// TIA Portal project "SSA-3GHz" (V15.1)

(* hardware
DEVICE "S7-1200"  S7-1200 Station
   slot 0: "Stand.sectionalRail35mmLength483mm_0"  S7-1200 Rack  Rack  V1.0
   slot 1: "S7-1200"  CPU 1215C DC/DC/DC  6ES7 215-1AG40-0XB0  V4.3
   slot 2: "AnalogInputSM12314AI_2"  6ES7 231-4HD32-0XB0  V2.0
   slot 3: "S7-1200analogInputSM1231RTD4AI_3"  SM 1231 AI4 x RTD  6ES7 231-5PD32-0XB0  V2.0
DEVICE "HMI_1"  KTP400 Basic PN
   slot 0: "HMI_1"  KTP400 Basic PN  6AV2 123-2DB03-0AX0  15.1.0.0
   slot 1: "HMI_RT_1"  KTP400 Basic PN  6AV2 123-2DB03-0AX0  15.1.0.0
   slot 5: "HMI_1.IE_CP_1"  PROFINET Interface  15.0.1.0
      slot 1: "PROFINET Interface_1"  PROFINET Interface
         slot 1: "Port_1"  Port
*)

// ===== PLC "S7-1200"  CPU 1215C DC/DC/DC =====

VAR_GLOBAL   // PLC tag table "Default tag table"
   "System_Byte" AT %MB1 : Byte;
   "FirstScan" AT %M1.0 : Bool;
   "DiagStatusUpdate" AT %M1.1 : Bool;
   "AlwaysTRUE" AT %M1.2 : Bool;
   "AlwaysFALSE" AT %M1.3 : Bool;
   "Clock_Byte" AT %MB0 : Byte;
   "Clock_10Hz" AT %M0.0 : Bool;
   "Clock_5Hz" AT %M0.1 : Bool;
   "Clock_2.5Hz" AT %M0.2 : Bool;
   "Clock_2Hz" AT %M0.3 : Bool;
   "Clock_1.25Hz" AT %M0.4 : Bool;
   "Clock_1Hz" AT %M0.5 : Bool;
   "Clock_0.625Hz" AT %M0.6 : Bool;
   "Clock_0.5Hz" AT %M0.7 : Bool;
   "MoveBlkStat" AT %MW100 : Int;
END_VAR

VAR_GLOBAL   // PLC tag table "Test tags"
   "Counter" AT %MD100 : UDInt;
   "TestBlink" AT %Q1.0 : Bool;
   "VisuTest" AT %MB104 : Byte;
END_VAR

VAR_GLOBAL   // PLC tag table "Analog I/O"
   "U_drain_RBK" AT %IW64 : Int;   // Drain voltage read-back
   "U_drain" AT %QW64 : Int;   // Drain voltage set-point
   "ADC0ch1" AT %IW66 : Int;   // Spare
   "U_gate" AT %QW66 : Int;   // Gate voltage set-point
   "Pfwd" AT %IW96 : Int;   // Forward power
   "Prev" AT %IW98 : Int;   // Reverse power
   "I_drain" AT %IW100 : Int;   // Drain current
   "U_gate_RBK" AT %IW102 : Int;   // Gate voltage read-back
   "TT001" AT %IW112 : Int;
   "TT002" AT %IW114 : Int;
   "TT003" AT %IW116 : Int;
   "TT004" AT %IW118 : Int;
END_VAR

VAR_GLOBAL   // PLC tag table "Digital I/O"
   "DutyCycOK" AT %I0.0 : Bool;   // Duty cycle OK
   "KeyIntlkOK" AT %I0.1 : Bool;   // Key interlock OK
   "ExtIntlkT1" AT %I0.2 : Bool;   // DC PS enable
   "ExtIntlkT3" AT %I0.3 : Bool;
   "PS_OK" AT %I0.4 : Bool;
   "CoolingWtrOK" AT %I0.5 : Bool;
   "KeyOK" AT %I0.6 : Bool;
   "FanOK" AT %I0.7 : Bool;
   "ExtIntlkOK" AT %I1.0 : Bool;
   "RFSwitchOn" AT %Q0.0 : Bool;   // Close RF switch
   "PScmdOn" AT %Q0.1 : Bool;   // Set PS On
   "SSA_OK" AT %Q0.2 : Bool;   // Solid State Amplifier OK
   "ResetOut" AT %Q0.3 : Bool;   // Reset the errors signal out
END_VAR

TYPE "DigitalIN"
   STRUCT
      DigitalIN : Struct
         PhysIn : Bool;   // Physical input
         NegLogic : Bool;   // 0 - positive lgic, 1 - negative logic
         Disabled : Bool;   // 0 - signal enabled, 1 - signal disabled (not used in process controll)
         Out : Bool;   // Logical value after taking into accout NegLogic setting
      END_STRUCT;
   END_STRUCT;
END_TYPE

TYPE "AnalogOUT"
   STRUCT
      AnalogOUT : Struct
         In : Real;
         Out : Int;
         VisuState : Byte;
         MINDAC : Int;
         MAXDAC : Int;
         MINEGU : Real;
         MAXEGU : Real;
      END_STRUCT;
   END_STRUCT;
END_TYPE

TYPE "AnalogIN"
   STRUCT
      AnalogIN : Struct
         In : Word;
         Out : Real;
         Low : Real;
         LoLo : Real;
         High : Real;
         HIHi : Real;
         VisuState : Byte;
         MINADC : Int;
         MAXADC : Int;
         MINEGU : Real;
         MAXEGU : Real;
      END_STRUCT;
   END_STRUCT;
END_TYPE

DATA_BLOCK "IEC_Counter_0_DB"   // DB5
{ S7_Optimized_Access := 'TRUE' }
AUTHOR : Simatic
FAMILY : IEC
NAME : UDCNTR
VERSION : 1.2
// stored: InstanceOfName IEC_UDCOUNTER
"IEC_UDCOUNTER"
BEGIN
END_DATA_BLOCK

DATA_BLOCK "ModbusData"   // DB100
{ S7_Optimized_Access := 'TRUE' }
VERSION : 0.1
   VAR
      serverData : Struct
         disconnect : Bool;
         ndr : Bool;
         dataRead : Bool;
         error : Bool;
         status : Word;
         statusSave : Word;
      END_STRUCT;
      connectParamServer : TCON_IP_v4;
   END_VAR
BEGIN
   connectParamServer.InterfaceId := 64;
   connectParamServer.ID := 16#1;
   connectParamServer.RemoteAddress.ADDR[1] := 0;
   connectParamServer.RemoteAddress.ADDR[2] := 0;
   connectParamServer.RemoteAddress.ADDR[3] := 0;
   connectParamServer.RemoteAddress.ADDR[4] := 0;
   connectParamServer.RemotePort := 0;
   connectParamServer.LocalPort := 502;
END_DATA_BLOCK

DATA_BLOCK "ModbusBuffer"   // DB101
{ S7_Optimized_Access := 'FALSE' }
VERSION : 0.1
   VAR
      BufferINOut : Struct
         LookupTable : Struct
            Pwr : Array[0..9] of Real;
            Ud : Array[0..9] of Real;
            Ug : Array[0..9] of Real;
         END_STRUCT;
         SetupData : Struct
            RemoteMode : Bool;   // When true- remote control only
            dBm_unit : Bool;   // When true - show power in dBm units
            NominalPower : Real := 100.0;   // Nominal Power
            NominalPower_dBm : Real;   // Nominal Pwr [dBm]
            UdSP : Real;   // Udrain set-point
            UgSP : Real;   // Ugate set-point
         END_STRUCT;
         Commands : Struct
            On : Bool;
            Off : Bool;
            Stdby : Bool;
            Reset : Bool;
         END_STRUCT;
         ADCdata : Struct
            Udrain : Real;
            Ugate : Real;
            Pfwd : Real;
            Prev : Real;
            Idrain : Real;
            spare : Real;
            TT01 : Real;
            TT02 : Real;
            TT03 : Real;
            TT04 : Real;
         END_STRUCT;
         CalculatedData : Struct
            Pfwd_dBm : Real;
            Prev_dBm : Real;
            spare : Array[0..9] of Int;
         END_STRUCT;
         StatusBits : Struct
            DutyCycOK : Bool;
            KeyIntlkOK : Bool;
            ExtIntlkT1 : Bool;
            ExtIntlkT3 : Bool;
            PS_OK : Bool;
            CoolingOK : Bool;
            FanOK : Bool;
            ExtIntlkOK : Bool;
            DutyCycOK_Ign : Bool;
            KeyIntlkOK_Ign : Bool;
            ExtIntlkT1_Ign : Bool;
            ExtIntlkT3_Ign : Bool;
            PS_OK_Ign : Bool;
            CoolingOK_Ign : Bool;
            FanOK_Ign : Bool;
            ExtIntlkOK_Ign : Bool;
         END_STRUCT;
      END_STRUCT;
   END_VAR
BEGIN
   BufferINOut.LookupTable.Pwr[0] := 10.0;
   BufferINOut.LookupTable.Pwr[1] := 20.0;
   BufferINOut.LookupTable.Pwr[2] := 50.0;
   BufferINOut.LookupTable.Pwr[3] := 100.0;
   BufferINOut.LookupTable.Pwr[4] := 200.0;
   BufferINOut.LookupTable.Pwr[5] := 300.0;
   BufferINOut.LookupTable.Pwr[6] := 400.0;
   BufferINOut.LookupTable.Ud[0] := 15.0;
   BufferINOut.LookupTable.Ud[1] := 17.0;
   BufferINOut.LookupTable.Ud[2] := 19.0;
   BufferINOut.LookupTable.Ud[3] := 22.0;
   BufferINOut.LookupTable.Ud[4] := 25.0;
   BufferINOut.LookupTable.Ud[5] := 30.0;
   BufferINOut.LookupTable.Ud[6] := 35.0;
   BufferINOut.LookupTable.Ug[0] := 1.5;
   BufferINOut.LookupTable.Ug[1] := 1.7;
   BufferINOut.LookupTable.Ug[2] := 1.9;
   BufferINOut.LookupTable.Ug[3] := 2.2;
   BufferINOut.LookupTable.Ug[4] := 2.5;
   BufferINOut.LookupTable.Ug[5] := 2.8;
   BufferINOut.LookupTable.Ug[6] := 3.0;
END_DATA_BLOCK

DATA_BLOCK "DigitalInputs"   // DB400
{ S7_Optimized_Access := 'TRUE' }
VERSION : 0.1
   VAR
      DutyCycOK : "DigitalIN";
      KeyIntlkOK : "DigitalIN";
      ExtIntlkT1 : "DigitalIN";
      ExtIntlkT3 : "DigitalIN";
      PS_OK : "DigitalIN";
      CoolingWtrOK : "DigitalIN";
      FanOK : "DigitalIN";
      ExtIntlkOK : "DigitalIN";
   END_VAR
BEGIN
   KeyIntlkOK.DigitalIN.Disabled := true;
   CoolingWtrOK.DigitalIN.Disabled := true;
   FanOK.DigitalIN.Disabled := true;
   ExtIntlkOK.DigitalIN.Disabled := true;
   PS_OK.DigitalIN.Disabled := true;
END_DATA_BLOCK

DATA_BLOCK "AnalogInputs"   // DB401
{ S7_Optimized_Access := 'TRUE' }
VERSION : 0.1
   VAR
      U_drain_RBK : "AnalogIN";
      U_gate_RBK : "AnalogIN";
      Pfwd : "AnalogIN";
      Prev : "AnalogIN";
      I_drain : "AnalogIN";
      ADC0ch1 : "AnalogIN";
      Pfwd_dBm : Real;
      Prev_dBm : Real;
   END_VAR
BEGIN
   U_drain_RBK.AnalogIN.MAXADC := 27648;
   U_gate_RBK.AnalogIN.MINADC := -27648;
   U_gate_RBK.AnalogIN.MAXADC := 27648;
   Pfwd.AnalogIN.MAXADC := 27648;
   Pfwd.AnalogIN.MAXEGU := 400.0;
   Prev.AnalogIN.MAXADC := 27648;
   Prev.AnalogIN.MAXEGU := 400.0;
   I_drain.AnalogIN.MAXADC := 27648;
   I_drain.AnalogIN.MAXEGU := 15.0;
   ADC0ch1.AnalogIN.MAXADC := 27648;
   ADC0ch1.AnalogIN.MAXEGU := 10.0;
   U_drain_RBK.AnalogIN.MAXEGU := 35.0;
   U_gate_RBK.AnalogIN.MAXEGU := 5.0;
   U_gate_RBK.AnalogIN.MINEGU := -5.0;
END_DATA_BLOCK

DATA_BLOCK "AnalogOutputs"   // DB402
{ S7_Optimized_Access := 'TRUE' }
VERSION : 0.1
   VAR
      U_drain : "AnalogOUT";
      U_gate : "AnalogOUT";
   END_VAR
BEGIN
   U_drain.AnalogOUT.MAXDAC := 27648;
   U_drain.AnalogOUT.MAXEGU := 35.0;
   U_gate.AnalogOUT.MAXDAC := 27648;
   U_gate.AnalogOUT.MAXEGU := 5.0;
   U_gate.AnalogOUT.MINEGU := 0.0;
END_DATA_BLOCK

DATA_BLOCK "DigitalOutputs"   // DB450
{ S7_Optimized_Access := 'TRUE' }
VERSION : 0.1
   VAR
      RF_Switch_ON : Bool;
      ResetCmd : Bool;
   END_VAR
BEGIN
END_DATA_BLOCK

DATA_BLOCK "LookupTable"   // DB500
{ S7_Optimized_Access := 'FALSE' }
VERSION : 0.1
   VAR
      Pwr : Array[0..9] of Real;
      Ud : Array[0..9] of Real;
      Ug : Array[0..9] of Real;
   END_VAR
BEGIN
   Pwr[0] := 10.0;
   Pwr[1] := 20.0;
   Pwr[2] := 50.0;
   Pwr[3] := 100.0;
   Pwr[4] := 200.0;
   Pwr[5] := 300.0;
   Pwr[6] := 400.0;
   Ud[0] := 15.0;
   Ud[1] := 17.0;
   Ud[2] := 19.0;
   Ud[3] := 22.0;
   Ud[4] := 25.0;
   Ud[5] := 30.0;
   Ud[6] := 35.0;
   Ug[0] := 1.5;
   Ug[1] := 1.7;
   Ug[2] := 1.9;
   Ug[3] := 2.2;
   Ug[4] := 2.5;
   Ug[5] := 2.8;
   Ug[6] := 3.0;
END_DATA_BLOCK

// folder: 5_T_CONFIG (S7-1200, S7-1500)

DATA_BLOCK "SLI_gDB_T_CONFIG_PLC"   // DB1
{ S7_Optimized_Access := 'TRUE' }
VERSION : 0.1
   VAR
      T_CONFIG : Struct   // Variables of T_CONFIG
         start : Bool;   // Set "start" to TRUE to configure the PROFINET interface.
         hwid : Hw_Interface := 64;   // Identification number of the PROFINET interface of the device (e. g. PROFINET interface of the CPU).
         busy : Bool;
         done : Bool;
         error : Bool;
         errorLocation : DWord;
         status : DWord;
         memErrStat : DWord;   // Saves the error status.
      END_STRUCT;
      configData : Struct   // Data to configure the PROFINET device.
         header : IF_CONF_Header;   // The header is used to define the number of system data types.
         deviceIP : IF_CONF_v4;   // Specifies the IP of the PROFINET device.
         deviceName : IF_CONF_NOS;   // Specifies the name of the PROFINET interface ("PROFINET device name").
      END_STRUCT;
   END_VAR
BEGIN
   configData.header.SubfieldCount := 2;   // 2: Indicates that two additional structures ("deviceIP" and "deviceName") are used below.
   configData.deviceName.Length := 11;   // Information on overall length of the structure (5 bytes for the device name "myplc" + 6 bytes for the parameters Id, Length and Mode)
   configData.deviceName.Mode := 1;   // 1: Permanent change of the device name in "myplc".
   configData.deviceName.NOS[1] := 'm';
   configData.deviceName.NOS[2] := 'y';
   configData.deviceName.NOS[3] := 'p';
   configData.deviceName.NOS[4] := 'l';
   configData.deviceName.NOS[5] := 'c';
   configData.deviceIP.Length := 18;   // Information on overall length of the structure (12 bytes for the device IP + 6 bytes for the parameters Id, Length and Mode)
   configData.deviceIP.Mode := 1;   // 1: Permanent change of the device IP.
   configData.deviceIP.InterfaceAddress.ADDR[1] := 192;
   configData.deviceIP.InterfaceAddress.ADDR[2] := 168;
   configData.deviceIP.InterfaceAddress.ADDR[3] := 0;
   configData.deviceIP.InterfaceAddress.ADDR[4] := 10;
   configData.deviceIP.SubnetMask.ADDR[1] := 255;
   configData.deviceIP.SubnetMask.ADDR[2] := 255;
   configData.deviceIP.SubnetMask.ADDR[3] := 255;
   configData.deviceIP.SubnetMask.ADDR[4] := 0;
   // configData.header.FieldType : Field type: Must always have the value "0".
   // configData.header.FieldId : Error ID: Must always have the value "0".
   // configData.deviceIP.Id : System data type ID. The start value of this parameter must not be changed.
   // configData.deviceIP.InterfaceAddress : IP connection data. IP address
   // configData.deviceIP.SubnetMask : IP connection data. Subnet mask
   // configData.deviceIP.DefaultRouter : IP connection data. Router address (optional)
   // configData.deviceName.Id : System data type ID. The start value of this parameter must not be changed.
   // configData.deviceName.NOS : Device name (1 character per byte)
END_DATA_BLOCK

DATA_BLOCK "SLI_gDB_T_CONFIG_HMI"   // DB4
{ S7_Optimized_Access := 'TRUE' }
VERSION : 0.1
   VAR
      T_CONFIG : Struct   // Variables of T_CONFIG
         start : Bool;   // Set "start" to TRUE to configure the PROFINET interface.
         hwid : Hw_Interface := 65;   // Identification number of the PROFINET interface of the device (e. g. PROFINET interface of the CPU).
         busy : Bool;
         done : Bool;
         error : Bool;
         errorLocation : DWord;
         status : DWord;
         memErrStat : DWord;   // Saves the error status.
      END_STRUCT;
      configData : Struct   // Data to configure the PROFINET device.
         header : IF_CONF_Header;   // The header is used to define the number of system data types.
         deviceIP : IF_CONF_v4;   // Specifies the IP of the PROFINET device.
         deviceName : IF_CONF_NOS;   // Specifies the name of the PROFINET interface ("PROFINET device name").
      END_STRUCT;
   END_VAR
BEGIN
   configData.header.SubfieldCount := 2;   // 2: Indicates that two additional structures ("deviceIP" and "deviceName") are used below.
   configData.deviceName.Length := 11;   // Information on overall length of the structure (5 bytes for the device name "myplc" + 6 bytes for the parameters Id, Length and Mode)
   configData.deviceName.Mode := 1;   // 1: Permanent change of the device name in "myplc".
   configData.deviceName.NOS[1] := 'm';
   configData.deviceName.NOS[2] := 'y';
   configData.deviceName.NOS[3] := 'h';
   configData.deviceName.NOS[4] := 'm';
   configData.deviceName.NOS[5] := 'i';
   configData.deviceIP.Length := 18;   // Information on overall length of the structure (12 bytes for the device IP + 6 bytes for the parameters Id, Length and Mode)
   configData.deviceIP.Mode := 1;   // 1: Permanent change of the device IP.
   configData.deviceIP.InterfaceAddress.ADDR[1] := 192;
   configData.deviceIP.InterfaceAddress.ADDR[2] := 168;
   configData.deviceIP.InterfaceAddress.ADDR[3] := 0;
   configData.deviceIP.InterfaceAddress.ADDR[4] := 11;
   configData.deviceIP.SubnetMask.ADDR[1] := 255;
   configData.deviceIP.SubnetMask.ADDR[2] := 255;
   configData.deviceIP.SubnetMask.ADDR[3] := 255;
   configData.deviceIP.SubnetMask.ADDR[4] := 0;
   // configData.header.FieldType : Field type: Must always have the value "0".
   // configData.header.FieldId : Error ID: Must always have the value "0".
   // configData.deviceIP.Id : System data type ID. The start value of this parameter must not be changed.
   // configData.deviceIP.InterfaceAddress : IP connection data. IP address
   // configData.deviceIP.SubnetMask : IP connection data. Subnet mask
   // configData.deviceIP.DefaultRouter : IP connection data. Router address (optional)
   // configData.deviceName.Id : System data type ID. The start value of this parameter must not be changed.
   // configData.deviceName.NOS : Device name (1 character per byte)
END_DATA_BLOCK

// folder: System blocks/Program resources

DATA_BLOCK "ResetCmdTimer"   // DB7
{ S7_Optimized_Access := 'TRUE' }
AUTHOR : Simatic
FAMILY : IEC
NAME : IEC_TMR
VERSION : 1.0
// stored: InstanceOfName IEC_TIMER
"IEC_TIMER"
BEGIN
END_DATA_BLOCK

// folder: (top level)

FUNCTION "Tests" : Void   // FC1, LAD
{ S7_Optimized_Access := 'TRUE' }
VERSION : 0.1
BEGIN

REGION Network 1
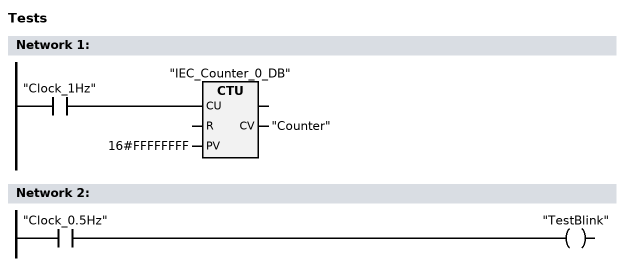
   "IEC_Counter_0_DB".CTU(CU := "Clock_1Hz", PV := 16#FFFFFFFF, CV => "Counter");
END_REGION

REGION Network 2
   RUNG wire#powerrail
      Contact( "Clock_0.5Hz" )
      Coil( "TestBlink" )
   END_RUNG
   // the same network as SCL:
   "TestBlink" := "Clock_0.5Hz";
END_REGION
END_FUNCTION

FUNCTION "Modbus2PLC" : Void   // FC10, LAD
{ S7_Optimized_Access := 'TRUE' }
VERSION : 0.1
BEGIN

REGION Network 1
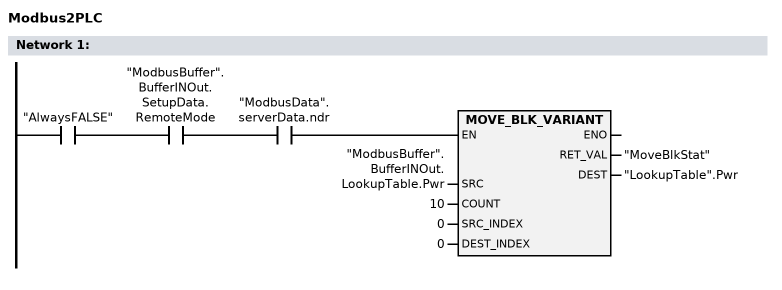
   IF "AlwaysFALSE" AND "ModbusBuffer".BufferINOut.SetupData.RemoteMode AND "ModbusData".serverData.ndr THEN
       "MoveBlkStat" := MOVE_BLK_VARIANT(SRC := "ModbusBuffer".BufferINOut.LookupTable.Pwr,
                               COUNT := 10,
                               SRC_INDEX := 0,
                               DEST_INDEX := 0,
                               DEST => "LookupTable".Pwr);
   END_IF;
END_REGION
END_FUNCTION

FUNCTION "PLC2Modbus" : Void   // FC11, LAD
{ S7_Optimized_Access := 'TRUE' }
VERSION : 0.1
BEGIN

REGION Network 1
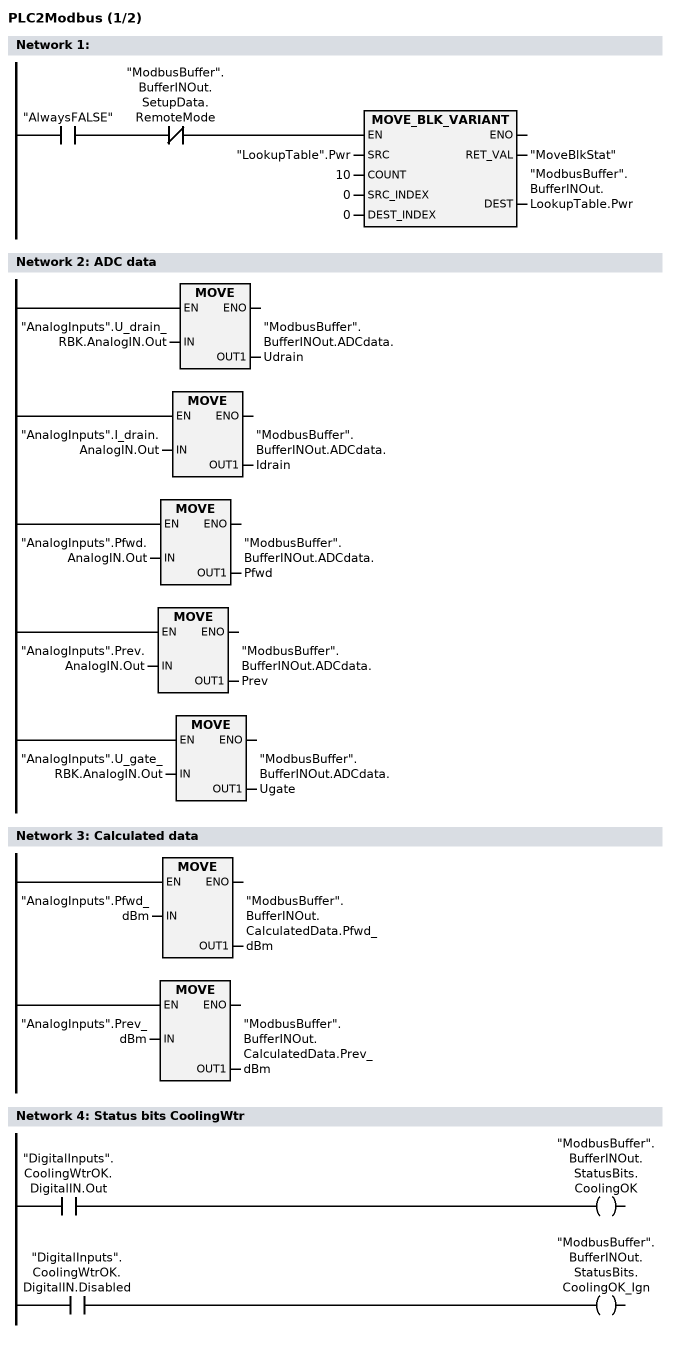
   IF "AlwaysFALSE" AND NOT "ModbusBuffer".BufferINOut.SetupData.RemoteMode THEN
       "MoveBlkStat" := MOVE_BLK_VARIANT(SRC := "LookupTable".Pwr,
                               COUNT := 10,
                               SRC_INDEX := 0,
                               DEST_INDEX := 0,
                               DEST => "ModbusBuffer".BufferINOut.LookupTable.Pwr);
   END_IF;
END_REGION

REGION Network 2: ADC data
   RUNG wire#powerrail
      Move(in := "AnalogInputs".U_drain_RBK.AnalogIN.Out, out1 => "ModbusBuffer".BufferINOut.ADCdata.Udrain)
   END_RUNG
   RUNG wire#powerrail
      Move(in := "AnalogInputs".I_drain.AnalogIN.Out, out1 => "ModbusBuffer".BufferINOut.ADCdata.Idrain)
   END_RUNG
   RUNG wire#powerrail
      Move(in := "AnalogInputs".Pfwd.AnalogIN.Out, out1 => "ModbusBuffer".BufferINOut.ADCdata.Pfwd)
   END_RUNG
   RUNG wire#powerrail
      Move(in := "AnalogInputs".Prev.AnalogIN.Out, out1 => "ModbusBuffer".BufferINOut.ADCdata.Prev)
   END_RUNG
   RUNG wire#powerrail
      Move(in := "AnalogInputs".U_gate_RBK.AnalogIN.Out, out1 => "ModbusBuffer".BufferINOut.ADCdata.Ugate)
   END_RUNG
   // the same network as SCL:
   "ModbusBuffer".BufferINOut.ADCdata.Udrain := "AnalogInputs".U_drain_RBK.AnalogIN.Out;
   "ModbusBuffer".BufferINOut.ADCdata.Idrain := "AnalogInputs".I_drain.AnalogIN.Out;
   "ModbusBuffer".BufferINOut.ADCdata.Pfwd := "AnalogInputs".Pfwd.AnalogIN.Out;
   "ModbusBuffer".BufferINOut.ADCdata.Prev := "AnalogInputs".Prev.AnalogIN.Out;
   "ModbusBuffer".BufferINOut.ADCdata.Ugate := "AnalogInputs".U_gate_RBK.AnalogIN.Out;
END_REGION

REGION Network 3: Calculated data
   RUNG wire#powerrail
      Move(in := "AnalogInputs".Pfwd_dBm, out1 => "ModbusBuffer".BufferINOut.CalculatedData.Pfwd_dBm)
   END_RUNG
   RUNG wire#powerrail
      Move(in := "AnalogInputs".Prev_dBm, out1 => "ModbusBuffer".BufferINOut.CalculatedData.Prev_dBm)
   END_RUNG
   // the same network as SCL:
   "ModbusBuffer".BufferINOut.CalculatedData.Pfwd_dBm := "AnalogInputs".Pfwd_dBm;
   "ModbusBuffer".BufferINOut.CalculatedData.Prev_dBm := "AnalogInputs".Prev_dBm;
END_REGION

REGION Network 4: Status bits CoolingWtr
   RUNG wire#powerrail
      Contact( "DigitalInputs".CoolingWtrOK.DigitalIN.Out )
      Coil( "ModbusBuffer".BufferINOut.StatusBits.CoolingOK )
   END_RUNG
   RUNG wire#powerrail
      Contact( "DigitalInputs".CoolingWtrOK.DigitalIN.Disabled )
      Coil( "ModbusBuffer".BufferINOut.StatusBits.CoolingOK_Ign )
   END_RUNG
   // the same network as SCL:
   "ModbusBuffer".BufferINOut.StatusBits.CoolingOK := "DigitalInputs".CoolingWtrOK.DigitalIN.Out;
   "ModbusBuffer".BufferINOut.StatusBits.CoolingOK_Ign := "DigitalInputs".CoolingWtrOK.DigitalIN.Disabled;
END_REGION

REGION Network 5: Status bits DutyCycOK
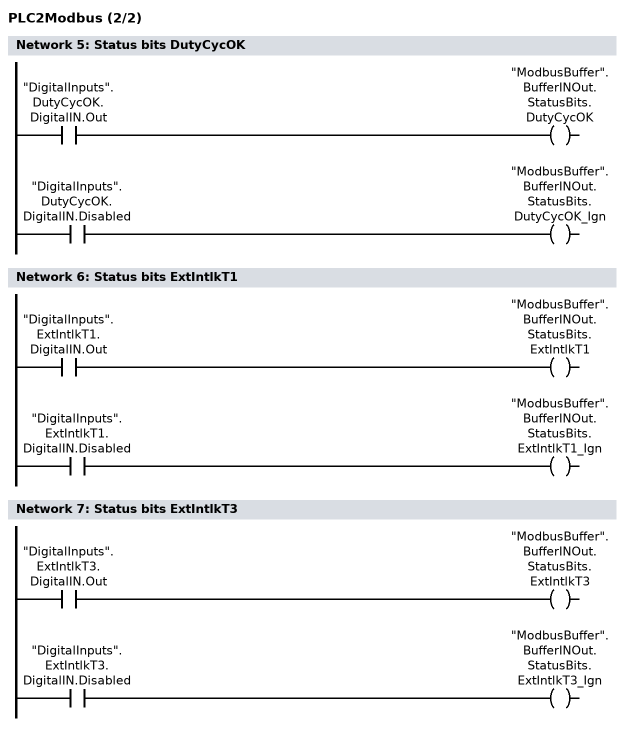
   RUNG wire#powerrail
      Contact( "DigitalInputs".DutyCycOK.DigitalIN.Out )
      Coil( "ModbusBuffer".BufferINOut.StatusBits.DutyCycOK )
   END_RUNG
   RUNG wire#powerrail
      Contact( "DigitalInputs".DutyCycOK.DigitalIN.Disabled )
      Coil( "ModbusBuffer".BufferINOut.StatusBits.DutyCycOK_Ign )
   END_RUNG
   // the same network as SCL:
   "ModbusBuffer".BufferINOut.StatusBits.DutyCycOK := "DigitalInputs".DutyCycOK.DigitalIN.Out;
   "ModbusBuffer".BufferINOut.StatusBits.DutyCycOK_Ign := "DigitalInputs".DutyCycOK.DigitalIN.Disabled;
END_REGION

REGION Network 6: Status bits ExtIntlkT1
   RUNG wire#powerrail
      Contact( "DigitalInputs".ExtIntlkT1.DigitalIN.Out )
      Coil( "ModbusBuffer".BufferINOut.StatusBits.ExtIntlkT1 )
   END_RUNG
   RUNG wire#powerrail
      Contact( "DigitalInputs".ExtIntlkT1.DigitalIN.Disabled )
      Coil( "ModbusBuffer".BufferINOut.StatusBits.ExtIntlkT1_Ign )
   END_RUNG
   // the same network as SCL:
   "ModbusBuffer".BufferINOut.StatusBits.ExtIntlkT1 := "DigitalInputs".ExtIntlkT1.DigitalIN.Out;
   "ModbusBuffer".BufferINOut.StatusBits.ExtIntlkT1_Ign := "DigitalInputs".ExtIntlkT1.DigitalIN.Disabled;
END_REGION

REGION Network 7: Status bits ExtIntlkT3
   RUNG wire#powerrail
      Contact( "DigitalInputs".ExtIntlkT3.DigitalIN.Out )
      Coil( "ModbusBuffer".BufferINOut.StatusBits.ExtIntlkT3 )
   END_RUNG
   RUNG wire#powerrail
      Contact( "DigitalInputs".ExtIntlkT3.DigitalIN.Disabled )
      Coil( "ModbusBuffer".BufferINOut.StatusBits.ExtIntlkT3_Ign )
   END_RUNG
   // the same network as SCL:
   "ModbusBuffer".BufferINOut.StatusBits.ExtIntlkT3 := "DigitalInputs".ExtIntlkT3.DigitalIN.Out;
   "ModbusBuffer".BufferINOut.StatusBits.ExtIntlkT3_Ign := "DigitalInputs".ExtIntlkT3.DigitalIN.Disabled;
END_REGION
END_FUNCTION

FUNCTION "Setup" : Void   // FC90, LAD
{ S7_Optimized_Access := 'TRUE' }
VERSION : 0.1
// Set-up PROFINET interfaces.
   VAR_TEMP
      done_PLC : Bool;
      done_HMI : Bool;
      errorLocation_PLC : DWord;
      errorLocation_HMI : DWord;
   END_VAR
BEGIN

REGION Network 1: Set "start" to TRUE to configure the PROFINET interface.
   // NOTE! Before using the example:
   // 
   // Condition:
   // 1) Open the device view of the CPU "> Properties > PROFINET interface > Ethernet addresses > PROFINET". 
   // 2) To set the device name: Activate the following options: 
   // - "IP address is set directly at the device". 
   // - "PROFINET device name is set directly at the device".
   // 
   // Regarding parameter INTERFACE ("hwid"):
   // - Change the value of "hwid" according to the identification number of the PROFINET interface of your local device (CPU). (Open "PLC tags > Show all tags > System constants. Look for a name like "<Local~PROFINET_interface_1>" with a Data type "Hw_Interface". The cell "value" contains the hwid.)
   // 
   // Info:
   // In the "header" (IF_CONF_HEADER):
   // - SubfieldCount = 2: Indicates that two additional structures ("deviceIP" and "deviceName") are used below.
   // 
   // In the structure "deviceIP" (system data type IF_CONF_v4):
   // - Lenght = 18: Information on overall length of the structure (12 bytes for the device IP + 6 bytes for the parameters Id, Length and Mode)
   // - Mode = 1: Permanent change of the device IP.
   // - InterfaceAddress, SubnetMask, DefaultRouter: IP connection data.
   // 
   // In the structure "deviceName" (system data type IF_CONF_NOS):
   // - Lenght = 11: Information on overall length of the structure (5 bytes for the device name "myplc" + 6 bytes for the parameters Id, Length and Mode)
   // - Mode = 1: Permanent change of the device name in "myplc".
   // - NOS[1] ... NOS[5]: Device name (1 character / byte)
   // 
   // Note: Instead of an absolute length, you can use the default start value (Lenght = 0) for a dynamic length.
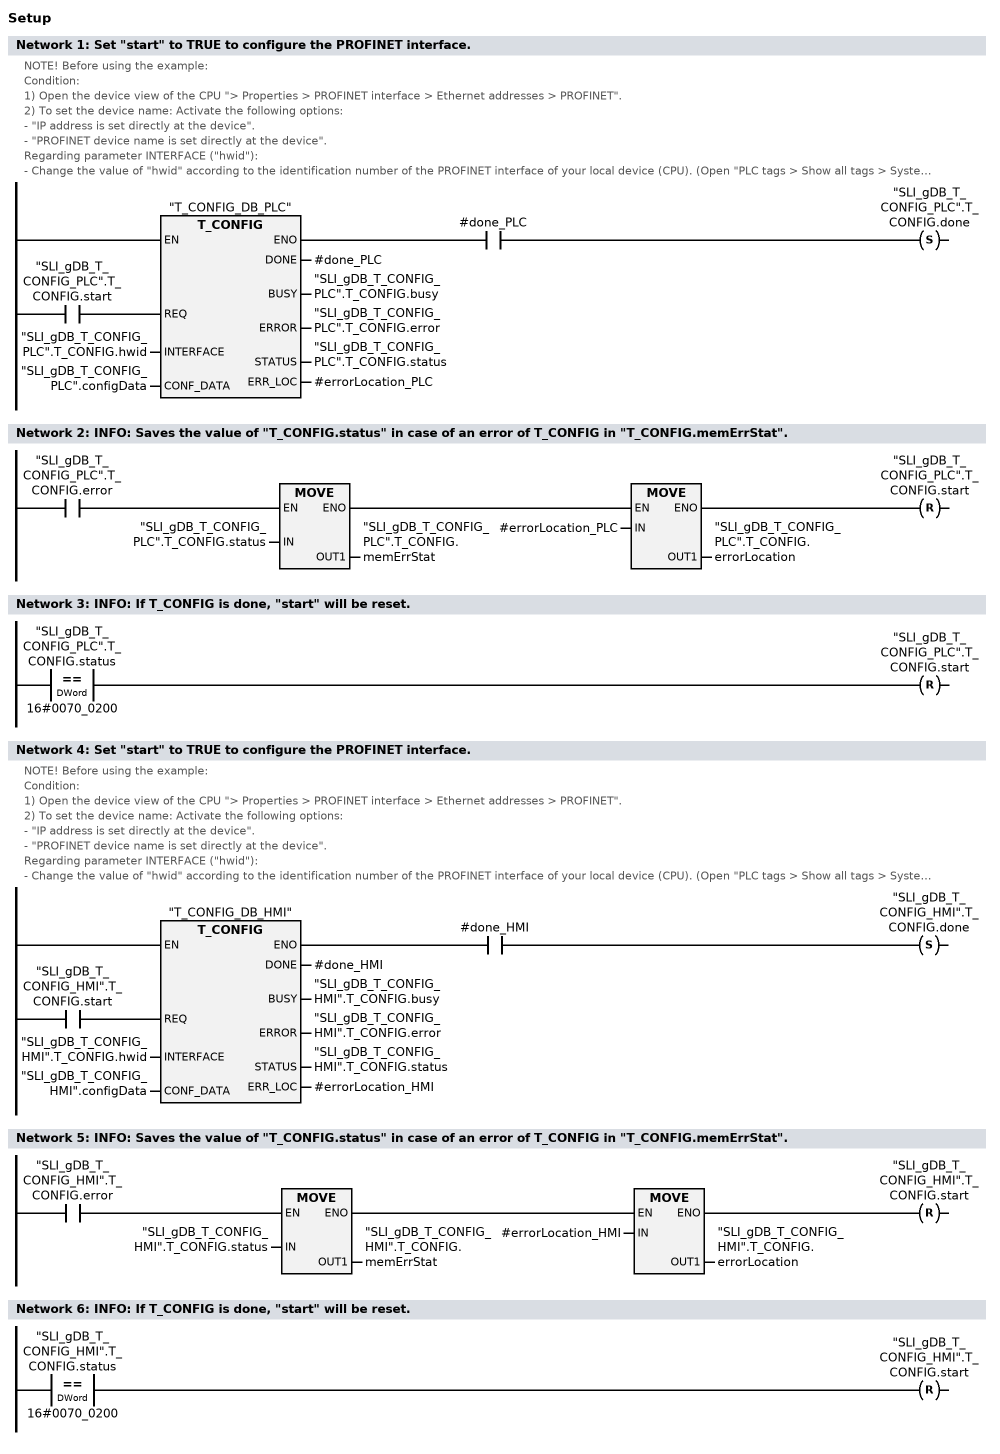
   // ENO of a box is taken as its EN; it also drops when the box reports an error
   "T_CONFIG_DB_PLC"(Req := "SLI_gDB_T_CONFIG_PLC".T_CONFIG.start,   // T_CONFIG
                     Interface := "SLI_gDB_T_CONFIG_PLC".T_CONFIG.hwid,
                     Conf_Data := "SLI_gDB_T_CONFIG_PLC".configData,
                     Done => #done_PLC,
                     Busy => "SLI_gDB_T_CONFIG_PLC".T_CONFIG.busy,
                     Error => "SLI_gDB_T_CONFIG_PLC".T_CONFIG.error,
                     Status => "SLI_gDB_T_CONFIG_PLC".T_CONFIG.status,
                     Err_Loc => #errorLocation_PLC);
   IF #done_PLC THEN "SLI_gDB_T_CONFIG_PLC".T_CONFIG.done := TRUE; END_IF;
END_REGION

REGION Network 2: INFO: Saves the value of "T_CONFIG.status" in case of an error of T_CONFIG in "T_CONFIG.memErrStat".
   RUNG wire#powerrail
      Contact( "SLI_gDB_T_CONFIG_PLC".T_CONFIG.error )
      Move(in := "SLI_gDB_T_CONFIG_PLC".T_CONFIG.status, out1 => "SLI_gDB_T_CONFIG_PLC".T_CONFIG.memErrStat)
      Move(in := #errorLocation_PLC, out1 => "SLI_gDB_T_CONFIG_PLC".T_CONFIG.errorLocation)
      R_Coil( "SLI_gDB_T_CONFIG_PLC".T_CONFIG.start )
   END_RUNG
   // the same network as SCL:
   IF "SLI_gDB_T_CONFIG_PLC".T_CONFIG.error THEN
       "SLI_gDB_T_CONFIG_PLC".T_CONFIG.memErrStat := "SLI_gDB_T_CONFIG_PLC".T_CONFIG.status;
       "SLI_gDB_T_CONFIG_PLC".T_CONFIG.errorLocation := #errorLocation_PLC;
       "SLI_gDB_T_CONFIG_PLC".T_CONFIG.start := FALSE;
   END_IF;
END_REGION

REGION Network 3: INFO: If T_CONFIG is done, "start" will be reset.
   RUNG wire#powerrail
      { S7_Templates := "SrcType := DWord" } EQ_Contact(in1 := "SLI_gDB_T_CONFIG_PLC".T_CONFIG.status, in2 := 16#0070_0200)
      R_Coil( "SLI_gDB_T_CONFIG_PLC".T_CONFIG.start )
   END_RUNG
   // the same network as SCL:
   IF "SLI_gDB_T_CONFIG_PLC".T_CONFIG.status = 16#0070_0200 THEN
       "SLI_gDB_T_CONFIG_PLC".T_CONFIG.start := FALSE;
   END_IF;
END_REGION

REGION Network 4: Set "start" to TRUE to configure the PROFINET interface.
   // NOTE! Before using the example:
   // 
   // Condition:
   // 1) Open the device view of the CPU "> Properties > PROFINET interface > Ethernet addresses > PROFINET". 
   // 2) To set the device name: Activate the following options: 
   // - "IP address is set directly at the device". 
   // - "PROFINET device name is set directly at the device".
   // 
   // Regarding parameter INTERFACE ("hwid"):
   // - Change the value of "hwid" according to the identification number of the PROFINET interface of your local device (CPU). (Open "PLC tags > Show all tags > System constants. Look for a name like "<Local~PROFINET_interface_1>" with a Data type "Hw_Interface". The cell "value" contains the hwid.)
   // 
   // Info:
   // In the "header" (IF_CONF_HEADER):
   // - SubfieldCount = 2: Indicates that two additional structures ("deviceIP" and "deviceName") are used below.
   // 
   // In the structure "deviceIP" (system data type IF_CONF_v4):
   // - Lenght = 18: Information on overall length of the structure (12 bytes for the device IP + 6 bytes for the parameters Id, Length and Mode)
   // - Mode = 1: Permanent change of the device IP.
   // - InterfaceAddress, SubnetMask, DefaultRouter: IP connection data.
   // 
   // In the structure "deviceName" (system data type IF_CONF_NOS):
   // - Lenght = 11: Information on overall length of the structure (5 bytes for the device name "myplc" + 6 bytes for the parameters Id, Length and Mode)
   // - Mode = 1: Permanent change of the device name in "myplc".
   // - NOS[1] ... NOS[5]: Device name (1 character / byte)
   // 
   // Note: Instead of an absolute length, you can use the default start value (Lenght = 0) for a dynamic length.
   // ENO of a box is taken as its EN; it also drops when the box reports an error
   "T_CONFIG_DB_HMI"(Req := "SLI_gDB_T_CONFIG_HMI".T_CONFIG.start,   // T_CONFIG
                     Interface := "SLI_gDB_T_CONFIG_HMI".T_CONFIG.hwid,
                     Conf_Data := "SLI_gDB_T_CONFIG_HMI".configData,
                     Done => #done_HMI,
                     Busy => "SLI_gDB_T_CONFIG_HMI".T_CONFIG.busy,
                     Error => "SLI_gDB_T_CONFIG_HMI".T_CONFIG.error,
                     Status => "SLI_gDB_T_CONFIG_HMI".T_CONFIG.status,
                     Err_Loc => #errorLocation_HMI);
   IF #done_HMI THEN "SLI_gDB_T_CONFIG_HMI".T_CONFIG.done := TRUE; END_IF;
END_REGION

REGION Network 5: INFO: Saves the value of "T_CONFIG.status" in case of an error of T_CONFIG in "T_CONFIG.memErrStat".
   RUNG wire#powerrail
      Contact( "SLI_gDB_T_CONFIG_HMI".T_CONFIG.error )
      Move(in := "SLI_gDB_T_CONFIG_HMI".T_CONFIG.status, out1 => "SLI_gDB_T_CONFIG_HMI".T_CONFIG.memErrStat)
      Move(in := #errorLocation_HMI, out1 => "SLI_gDB_T_CONFIG_HMI".T_CONFIG.errorLocation)
      R_Coil( "SLI_gDB_T_CONFIG_HMI".T_CONFIG.start )
   END_RUNG
   // the same network as SCL:
   IF "SLI_gDB_T_CONFIG_HMI".T_CONFIG.error THEN
       "SLI_gDB_T_CONFIG_HMI".T_CONFIG.memErrStat := "SLI_gDB_T_CONFIG_HMI".T_CONFIG.status;
       "SLI_gDB_T_CONFIG_HMI".T_CONFIG.errorLocation := #errorLocation_HMI;
       "SLI_gDB_T_CONFIG_HMI".T_CONFIG.start := FALSE;
   END_IF;
END_REGION

REGION Network 6: INFO: If T_CONFIG is done, "start" will be reset.
   RUNG wire#powerrail
      { S7_Templates := "SrcType := DWord" } EQ_Contact(in1 := "SLI_gDB_T_CONFIG_HMI".T_CONFIG.status, in2 := 16#0070_0200)
      R_Coil( "SLI_gDB_T_CONFIG_HMI".T_CONFIG.start )
   END_RUNG
   // the same network as SCL:
   IF "SLI_gDB_T_CONFIG_HMI".T_CONFIG.status = 16#0070_0200 THEN
       "SLI_gDB_T_CONFIG_HMI".T_CONFIG.start := FALSE;
   END_IF;
END_REGION
END_FUNCTION

FUNCTION "ProcessDI" : Void   // FC400, LAD
{ S7_Optimized_Access := 'TRUE' }
VERSION : 0.1
BEGIN

REGION Network 1: DutyCycOK
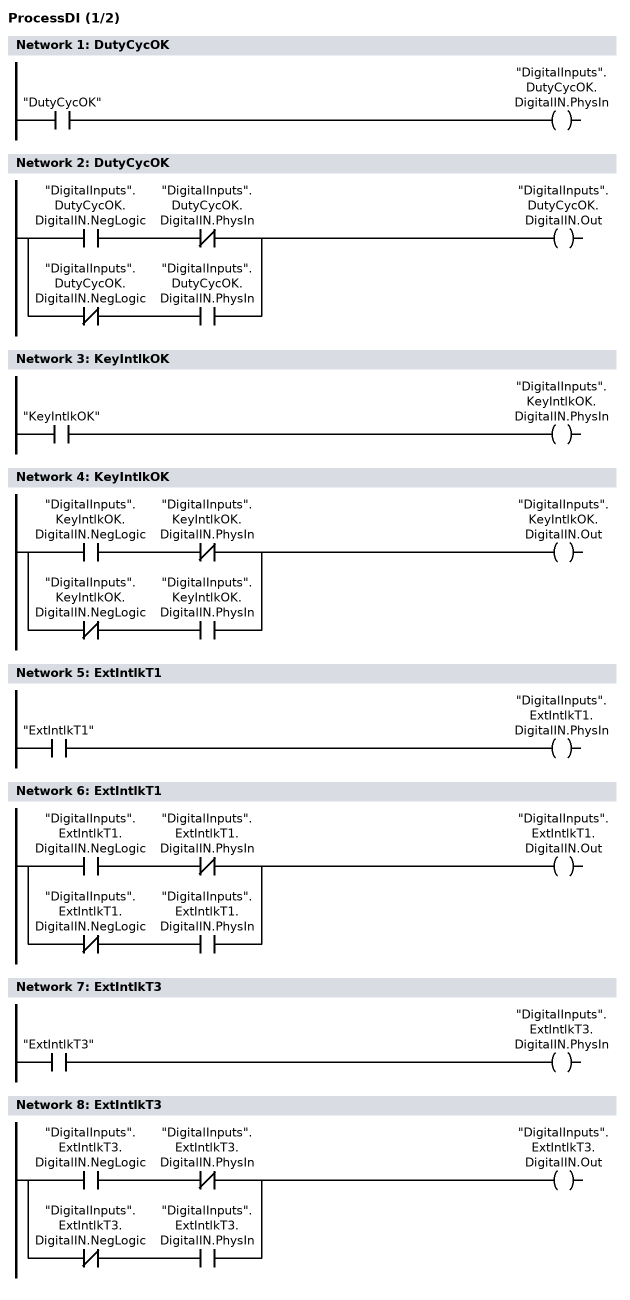
   RUNG wire#powerrail
      Contact( "DutyCycOK" )
      Coil( "DigitalInputs".DutyCycOK.DigitalIN.PhysIn )
   END_RUNG
   // the same network as SCL:
   "DigitalInputs".DutyCycOK.DigitalIN.PhysIn := "DutyCycOK";
END_REGION

REGION Network 2: DutyCycOK
   RUNG wire#powerrail
      Contact( "DigitalInputs".DutyCycOK.DigitalIN.NegLogic )
      I_Contact( "DigitalInputs".DutyCycOK.DigitalIN.PhysIn )
      wire#w1
      Coil( "DigitalInputs".DutyCycOK.DigitalIN.Out )
   END_RUNG
   RUNG wire#powerrail
      I_Contact( "DigitalInputs".DutyCycOK.DigitalIN.NegLogic )
      Contact( "DigitalInputs".DutyCycOK.DigitalIN.PhysIn )
   END_RUNG wire#w1
   // the same network as SCL:
   "DigitalInputs".DutyCycOK.DigitalIN.Out := ("DigitalInputs".DutyCycOK.DigitalIN.NegLogic AND NOT "DigitalInputs".DutyCycOK.DigitalIN.PhysIn) OR (NOT "DigitalInputs".DutyCycOK.DigitalIN.NegLogic AND "DigitalInputs".DutyCycOK.DigitalIN.PhysIn);
END_REGION

REGION Network 3: KeyIntlkOK
   RUNG wire#powerrail
      Contact( "KeyIntlkOK" )
      Coil( "DigitalInputs".KeyIntlkOK.DigitalIN.PhysIn )
   END_RUNG
   // the same network as SCL:
   "DigitalInputs".KeyIntlkOK.DigitalIN.PhysIn := "KeyIntlkOK";
END_REGION

REGION Network 4: KeyIntlkOK
   RUNG wire#powerrail
      Contact( "DigitalInputs".KeyIntlkOK.DigitalIN.NegLogic )
      I_Contact( "DigitalInputs".KeyIntlkOK.DigitalIN.PhysIn )
      wire#w1
      Coil( "DigitalInputs".KeyIntlkOK.DigitalIN.Out )
   END_RUNG
   RUNG wire#powerrail
      I_Contact( "DigitalInputs".KeyIntlkOK.DigitalIN.NegLogic )
      Contact( "DigitalInputs".KeyIntlkOK.DigitalIN.PhysIn )
   END_RUNG wire#w1
   // the same network as SCL:
   "DigitalInputs".KeyIntlkOK.DigitalIN.Out := ("DigitalInputs".KeyIntlkOK.DigitalIN.NegLogic AND NOT "DigitalInputs".KeyIntlkOK.DigitalIN.PhysIn) OR (NOT "DigitalInputs".KeyIntlkOK.DigitalIN.NegLogic AND "DigitalInputs".KeyIntlkOK.DigitalIN.PhysIn);
END_REGION

REGION Network 5: ExtIntlkT1
   RUNG wire#powerrail
      Contact( "ExtIntlkT1" )
      Coil( "DigitalInputs".ExtIntlkT1.DigitalIN.PhysIn )
   END_RUNG
   // the same network as SCL:
   "DigitalInputs".ExtIntlkT1.DigitalIN.PhysIn := "ExtIntlkT1";
END_REGION

REGION Network 6: ExtIntlkT1
   RUNG wire#powerrail
      Contact( "DigitalInputs".ExtIntlkT1.DigitalIN.NegLogic )
      I_Contact( "DigitalInputs".ExtIntlkT1.DigitalIN.PhysIn )
      wire#w1
      Coil( "DigitalInputs".ExtIntlkT1.DigitalIN.Out )
   END_RUNG
   RUNG wire#powerrail
      I_Contact( "DigitalInputs".ExtIntlkT1.DigitalIN.NegLogic )
      Contact( "DigitalInputs".ExtIntlkT1.DigitalIN.PhysIn )
   END_RUNG wire#w1
   // the same network as SCL:
   "DigitalInputs".ExtIntlkT1.DigitalIN.Out := ("DigitalInputs".ExtIntlkT1.DigitalIN.NegLogic AND NOT "DigitalInputs".ExtIntlkT1.DigitalIN.PhysIn) OR (NOT "DigitalInputs".ExtIntlkT1.DigitalIN.NegLogic AND "DigitalInputs".ExtIntlkT1.DigitalIN.PhysIn);
END_REGION

REGION Network 7: ExtIntlkT3
   RUNG wire#powerrail
      Contact( "ExtIntlkT3" )
      Coil( "DigitalInputs".ExtIntlkT3.DigitalIN.PhysIn )
   END_RUNG
   // the same network as SCL:
   "DigitalInputs".ExtIntlkT3.DigitalIN.PhysIn := "ExtIntlkT3";
END_REGION

REGION Network 8: ExtIntlkT3
   RUNG wire#powerrail
      Contact( "DigitalInputs".ExtIntlkT3.DigitalIN.NegLogic )
      I_Contact( "DigitalInputs".ExtIntlkT3.DigitalIN.PhysIn )
      wire#w1
      Coil( "DigitalInputs".ExtIntlkT3.DigitalIN.Out )
   END_RUNG
   RUNG wire#powerrail
      I_Contact( "DigitalInputs".ExtIntlkT3.DigitalIN.NegLogic )
      Contact( "DigitalInputs".ExtIntlkT3.DigitalIN.PhysIn )
   END_RUNG wire#w1
   // the same network as SCL:
   "DigitalInputs".ExtIntlkT3.DigitalIN.Out := ("DigitalInputs".ExtIntlkT3.DigitalIN.NegLogic AND NOT "DigitalInputs".ExtIntlkT3.DigitalIN.PhysIn) OR (NOT "DigitalInputs".ExtIntlkT3.DigitalIN.NegLogic AND "DigitalInputs".ExtIntlkT3.DigitalIN.PhysIn);
END_REGION

REGION Network 9: PS_OK
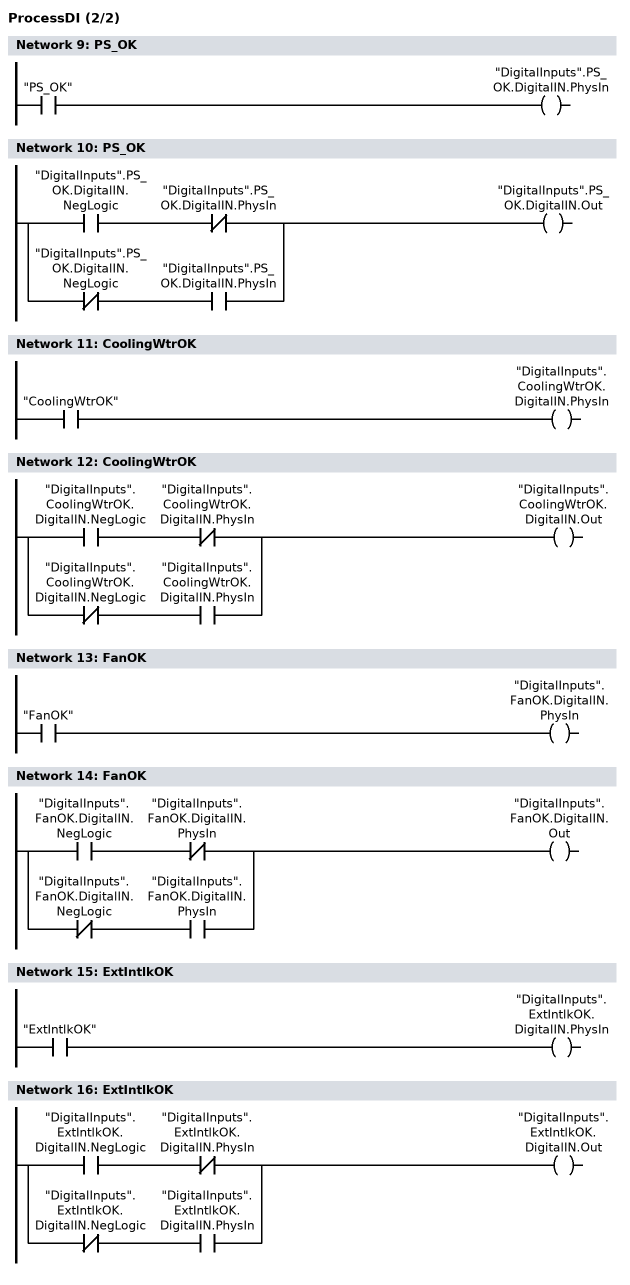
   RUNG wire#powerrail
      Contact( "PS_OK" )
      Coil( "DigitalInputs".PS_OK.DigitalIN.PhysIn )
   END_RUNG
   // the same network as SCL:
   "DigitalInputs".PS_OK.DigitalIN.PhysIn := "PS_OK";
END_REGION

REGION Network 10: PS_OK
   RUNG wire#powerrail
      Contact( "DigitalInputs".PS_OK.DigitalIN.NegLogic )
      I_Contact( "DigitalInputs".PS_OK.DigitalIN.PhysIn )
      wire#w1
      Coil( "DigitalInputs".PS_OK.DigitalIN.Out )
   END_RUNG
   RUNG wire#powerrail
      I_Contact( "DigitalInputs".PS_OK.DigitalIN.NegLogic )
      Contact( "DigitalInputs".PS_OK.DigitalIN.PhysIn )
   END_RUNG wire#w1
   // the same network as SCL:
   "DigitalInputs".PS_OK.DigitalIN.Out := ("DigitalInputs".PS_OK.DigitalIN.NegLogic AND NOT "DigitalInputs".PS_OK.DigitalIN.PhysIn) OR (NOT "DigitalInputs".PS_OK.DigitalIN.NegLogic AND "DigitalInputs".PS_OK.DigitalIN.PhysIn);
END_REGION

REGION Network 11: CoolingWtrOK
   RUNG wire#powerrail
      Contact( "CoolingWtrOK" )
      Coil( "DigitalInputs".CoolingWtrOK.DigitalIN.PhysIn )
   END_RUNG
   // the same network as SCL:
   "DigitalInputs".CoolingWtrOK.DigitalIN.PhysIn := "CoolingWtrOK";
END_REGION
